   "Carrier_74_Status.7" AT %I4050.7 : Bool;   // CARRIER FAULT
   "Carrier_74_Status.8" AT %I4051.0 : Bool;   // CRASH DETECT TRIPPED
   "Carrier_74_Status.9" AT %I4051.1 : Bool;
   "Carrier_74_Status.10" AT %I4051.2 : Bool;
   "Carrier_74_Status.11" AT %I4051.3 : Bool;
   "Carrier_74_Status.12" AT %I4051.4 : Bool;
   "Carrier_74_Status.13" AT %I4051.5 : Bool;
   "Carrier_74_Status.14" AT %I4051.6 : Bool;
   "Carrier_74_Status.15" AT %I4051.7 : Bool;
   "Carrier_74_SDCFaultCode" AT %IW4052 : Word;   // SDC FAULT CODE
   "Carrier_74_CarrierPosition" AT %ID4054 : DWord;   // CARRIER POSITION
   "Carrier_74_CarrierNumber" AT %IW4058 : Word;   // CARRIER NUMBER
   "Carrier_74_G120DControlWord" AT %IW4060 : Word;   // G120D_STW1_CONTROL
   "Carrier_74_G120DControlWord.0" AT %I4060.0 : Bool;   // Bit_00_ON
   "Carrier_74_G120DControlWord.1" AT %I4060.1 : Bool;   // Bit_01_AUS2_INH
   "Carrier_74_G120DControlWord.2" AT %I4060.2 : Bool;   // Bit_02_AUS3_STOP
   "Carrier_74_G120DControlWord.3" AT %I4060.3 : Bool;   // Bit_03_EN
   "Carrier_74_G120DControlWord.4" AT %I4060.4 : Bool;   // Bit_04_EN_RAMP
   "Carrier_74_G120DControlWord.5" AT %I4060.5 : Bool;   // Bit_05_START_RAMP
   "Carrier_74_G120DControlWord.6" AT %I4060.6 : Bool;   // Bit_06_SETPOINT
   "Carrier_74_G120DControlWord.7" AT %I4060.7 : Bool;   // Bit_07_RESET
   "Carrier_74_G120DControlWord.8" AT %I4061.0 : Bool;   // Bit_08_JOG_R
   "Carrier_74_G120DControlWord.9" AT %I4061.1 : Bool;   // Bit_09_JOG_L
   "Carrier_74_G120DControlWord.10" AT %I4061.2 : Bool;   // Bit_10_CONTR_PLC
   "Carrier_74_G120DControlWord.11" AT %I4061.3 : Bool;   // Bit_11_REVERSE
   "Carrier_74_G120DControlWord.12" AT %I4061.4 : Bool;   // Bit_12_BRAKE_RELEASE
   "Carrier_74_G120DControlWord.13" AT %I4061.5 : Bool;   // Bit_13_DDS
   "Carrier_74_G120DControlWord.14" AT %I4061.6 : Bool;   // Bit_14_DO0
   "Carrier_74_G120DControlWord.15" AT %I4061.7 : Bool;   // Bit_15_DO1
   "Carrier_74_G120DStatusWord" AT %IW4062 : Word;   // G120D_ZSW1_STATUS
   "Carrier_74_G120DStatusWord.0" AT %I4062.0 : Bool;   // Bit_00_READY_RUN
   "Carrier_74_G120DStatusWord.1" AT %I4062.1 : Bool;   // Bit_01_READY_ON
   "Carrier_74_G120DStatusWord.2" AT %I4062.2 : Bool;   // Bit_02_ENABLE
   "Carrier_74_G120DStatusWord.3" AT %I4062.3 : Bool;   // Bit_03_FAULT
   "Carrier_74_G120DStatusWord.4" AT %I4062.4 : Bool;   // Bit_04_OFF2
   "Carrier_74_G120DStatusWord.5" AT %I4062.5 : Bool;   // Bit_05_OFF3
   "Carrier_74_G120DStatusWord.6" AT %I4062.6 : Bool;   // Bit_06_LOCK_OUT
   "Carrier_74_G120DStatusWord.7" AT %I4062.7 : Bool;   // Bit_07_WARN
   "Carrier_74_G120DStatusWord.8" AT %I4063.0 : Bool;   // Bit_08_NO_DEVIATION
   "Carrier_74_G120DStatusWord.9" AT %I4063.1 : Bool;   // Bit_09_CONTR_PLC
   "Carrier_74_G120DStatusWord.10" AT %I4063.2 : Bool;   // Bit_10_F_MAX
   "Carrier_74_G120DStatusWord.11" AT %I4063.3 : Bool;   // Bit_11_LIMIT_REACHED
   "Carrier_74_G120DStatusWord.12" AT %I4063.4 : Bool;   // Bit_12_BRAKE_OPEN
   "Carrier_74_G120DStatusWord.13" AT %I4063.5 : Bool;   // Bit_13_NO_OVERTEMP
   "Carrier_74_G120DStatusWord.14" AT %I4063.6 : Bool;   // Bit_14_CW_CCW
   "Carrier_74_G120DStatusWord.15" AT %I4063.7 : Bool;   // Bit_15_OVERL
   "Carrier_74_Slot2_Input" AT %IW4064 : Word;   // SLOT 2 INPUT WORD
   "Carrier_74_CrashDetectSW" AT %I4064.0 : Bool;   // CRASH DETECT SW
   "Carrier_74_SpareSafetyInput(2_1)" AT %I4064.1 : Bool;   // SPARE SAFETY INPUT
   "Carrier_74_SpareSafetyInput(2_2)" AT %I4064.2 : Bool;   // SPARE SAFETY INPUT
   "Carrier_74_SpareSafetyInput(2_3)" AT %I4064.3 : Bool;   // SPARE SAFETY INPUT
   "Carrier_74_SpareSafetyInput(2_4)" AT %I4064.4 : Bool;   // SPARE SAFETY INPUT
   "Carrier_74_SpareSafetyInput(2_5)" AT %I4064.5 : Bool;   // SPARE SAFETY INPUT
   "Carrier_74_SpareSafetyInput(2_6)" AT %I4064.6 : Bool;   // SPARE SAFETY INPUT
   "Carrier_74_SpareSafetyInput(2_7)" AT %I4064.7 : Bool;   // SPARE SAFETY INPUT
   "Carrier_74_Slot3_SafetyOutput" AT %IW4065 : Word;   // SLOT 3 SAFETY OUTPUT WORD
   "Carrier_74_Crash_Detect_OK" AT %I4065.0 : Bool;   // CARRIER CRASH DETECT
   "Carrier_74_SpareSafetyOutput(3_1)" AT %I4065.1 : Bool;   // SPARE SAFETY OUTPUT
   "Carrier_74_SpareSafetyOutput(3_2)" AT %I4065.2 : Bool;   // SPARE SAFETY OUTPUT
   "Carrier_74_SpareSafetyOutput(3_3)" AT %I4065.3 : Bool;   // SPARE SAFETY OUTPUT
   "Carrier_74_SpareSafetyOutput(3_4)" AT %I4065.4 : Bool;   // SPARE SAFETY OUTPUT
   "Carrier_74_SpareSafetyOutput(3_5)" AT %I4065.5 : Bool;   // SPARE SAFETY OUTPUT
   "Carrier_74_SpareSafetyOutput(3_6)" AT %I4065.6 : Bool;   // SPARE SAFETY OUTPUT
   "Carrier_74_SpareSafetyOutput(3_7)" AT %I4065.7 : Bool;   // SPARE SAFETY OUTPUT
   "Carrier_74_Slot4_Input" AT %IW4066 : Word;   // SLOT 4 INPUT WORD
   "Carrier_74_480VPowerOn_MDCB1" AT %I4066.0 : Bool;   // 480 VAC POWER ON MDCB 1
   "Carrier_74_SpareInput(4_1)" AT %I4066.1 : Bool;   // SPARE INPUT
   "Carrier_74_SpareInput(4_2)" AT %I4066.2 : Bool;   // SPARE INPUT
   "Carrier_74_SitopSelectStatus" AT %I4066.3 : Bool;   // SITOP SELECT STATUS
   "Carrier_74_DCsupplyOnPSCB2" AT %I4066.4 : Bool;   // DC SUPPLY ON PSCB 2
   "Carrier_74_SpareInput(4_5)" AT %I4066.5 : Bool;   // SPARE INPUT
   "Carrier_74_SpareInput(4_6)" AT %I4066.6 : Bool;   // SPARE INPUT
   "Carrier_74_SpareInput(4_7)" AT %I4066.7 : Bool;   // SPARE INPUT
   "Carrier_74_PB1_ProdHoldLH" AT %I4067.0 : Bool;   // PB 1 PRODUCTION HOLD LH
   "Carrier_74_PB2_ResetLH" AT %I4067.1 : Bool;   // PB 2 RESET LH
   "Carrier_74_PB3_ProdHoldRH" AT %I4067.2 : Bool;   // PB 3 PRODUCTION HOLD RH
   "Carrier_74_PB4_ResetRH" AT %I4067.3 : Bool;   // PB 4 RESET RH
   "Carrier_74_SpareInput(4_14)" AT %I4067.4 : Bool;   // SPARE INPUT
   "Carrier_74_SpareInput(4_15)" AT %I4067.5 : Bool;   // SPARE INPUT
   "Carrier_74_SpareInput(4_16)" AT %I4067.6 : Bool;   // SPARE INPUT
   "Carrier_74_SpareInput(4_17)" AT %I4067.7 : Bool;   // SPARE INPUT
   "Carrier_74_Slot5_Output" AT %IW4068 : Word;   // SLOT 5 OUTPUT WORD
   "Carrier_74_IRD400_HMI_24VDC_ENABLE" AT %I4068.0 : Bool;   // IRD 400 PANEL HMI 24V DC POWER
   "Carrier_74_FaultLight_LH" AT %I4068.1 : Bool;   // FAULT LIGHT LH
   "Carrier_74_RunLight_LH" AT %I4068.2 : Bool;   // RUN LIGHT LH
   "Carrier_74_FaultLight_RH" AT %I4068.3 : Bool;   // FAULT LIGHT RH
   "Carrier_74_RunLight_RH" AT %I4068.4 : Bool;   // RUN LIGHT RH
   "Carrier_74_SpareOutput(5_5)" AT %I4068.5 : Bool;   // SPARE OUTPUT
   "Carrier_74_SpareOutput(5_6)" AT %I4068.6 : Bool;   // SPARE OUTPUT
   "Carrier_74_SpareOutput(5_7)" AT %I4068.7 : Bool;   // SPARE OUTPUT
   "Carrier_74_ActualSpeed" AT %IW4070 : Word;   // ACTUAL SPEED
   "Carrier_74_CarrierDriveAlarm" AT %IW4072 : Word;   // CARRIER DRIVE ALARM
   "Carrier_74_CarrierDriveWarning" AT %IW4074 : Word;   // CARRIER DRIVE WARNING
   "Carrier_75_Status" AT %IW4100 : Word;   // CARRIER STATUS WORD
   "Carrier_75_Status.0" AT %I4100.0 : Bool;   // HEARTBEAT
   "Carrier_75_Status.1" AT %I4100.1 : Bool;   // MANUAL
   "Carrier_75_Status.2" AT %I4100.2 : Bool;   // IN_AUTO
   "Carrier_75_Status.3" AT %I4100.3 : Bool;   // POSITIONING_COMPLETE
   "Carrier_75_Status.4" AT %I4100.4 : Bool;   // PRODUCTION HOLD
   "Carrier_75_Status.5" AT %I4100.5 : Bool;   // CARRIER MOVING FORWARD
   "Carrier_75_Status.6" AT %I4100.6 : Bool;   // CARRIER MOVING REVERSE
   "Carrier_75_Status.7" AT %I4100.7 : Bool;   // CARRIER FAULT
   "Carrier_75_Status.8" AT %I4101.0 : Bool;   // CRASH DETECT TRIPPED
   "Carrier_75_Status.9" AT %I4101.1 : Bool;
   "Carrier_75_Status.10" AT %I4101.2 : Bool;
   "Carrier_75_Status.11" AT %I4101.3 : Bool;
   "Carrier_75_Status.12" AT %I4101.4 : Bool;
   "Carrier_75_Status.13" AT %I4101.5 : Bool;
   "Carrier_75_Status.14" AT %I4101.6 : Bool;
   "Carrier_75_Status.15" AT %I4101.7 : Bool;
   "Carrier_75_SDCFaultCode" AT %IW4102 : Word;   // SDC FAULT CODE
   "Carrier_75_CarrierPosition" AT %ID4104 : DWord;   // CARRIER POSITION
   "Carrier_75_CarrierNumber" AT %IW4108 : Word;   // CARRIER NUMBER
   "Carrier_75_G120DControlWord" AT %IW4110 : Word;   // G120D_STW1_CONTROL
   "Carrier_75_G120DControlWord.0" AT %I4110.0 : Bool;   // Bit_00_ON
   "Carrier_75_G120DControlWord.1" AT %I4110.1 : Bool;   // Bit_01_AUS2_INH
   "Carrier_75_G120DControlWord.2" AT %I4110.2 : Bool;   // Bit_02_AUS3_STOP
   "Carrier_75_G120DControlWord.3" AT %I4110.3 : Bool;   // Bit_03_EN
   "Carrier_75_G120DControlWord.4" AT %I4110.4 : Bool;   // Bit_04_EN_RAMP
   "Carrier_75_G120DControlWord.5" AT %I4110.5 : Bool;   // Bit_05_START_RAMP
   "Carrier_75_G120DControlWord.6" AT %I4110.6 : Bool;   // Bit_06_SETPOINT
   "Carrier_75_G120DControlWord.7" AT %I4110.7 : Bool;   // Bit_07_RESET
   "Carrier_75_G120DControlWord.8" AT %I4111.0 : Bool;   // Bit_08_JOG_R
   "Carrier_75_G120DControlWord.9" AT %I4111.1 : Bool;   // Bit_09_JOG_L
   "Carrier_75_G120DControlWord.10" AT %I4111.2 : Bool;   // Bit_10_CONTR_PLC
   "Carrier_75_G120DControlWord.11" AT %I4111.3 : Bool;   // Bit_11_REVERSE
   "Carrier_75_G120DControlWord.12" AT %I4111.4 : Bool;   // Bit_12_BRAKE_RELEASE
   "Carrier_75_G120DControlWord.13" AT %I4111.5 : Bool;   // Bit_13_DDS
   "Carrier_75_G120DControlWord.14" AT %I4111.6 : Bool;   // Bit_14_DO0
   "Carrier_75_G120DControlWord.15" AT %I4111.7 : Bool;   // Bit_15_DO1
   "Carrier_75_G120DStatusWord" AT %IW4112 : Word;   // G120D_ZSW1_STATUS
   "Carrier_75_G120DStatusWord.0" AT %I4112.0 : Bool;   // Bit_00_READY_RUN
   "Carrier_75_G120DStatusWord.1" AT %I4112.1 : Bool;   // Bit_01_READY_ON
   "Carrier_75_G120DStatusWord.2" AT %I4112.2 : Bool;   // Bit_02_ENABLE
   "Carrier_75_G120DStatusWord.3" AT %I4112.3 : Bool;   // Bit_03_FAULT
   "Carrier_75_G120DStatusWord.4" AT %I4112.4 : Bool;   // Bit_04_OFF2
   "Carrier_75_G120DStatusWord.5" AT %I4112.5 : Bool;   // Bit_05_OFF3
   "Carrier_75_G120DStatusWord.6" AT %I4112.6 : Bool;   // Bit_06_LOCK_OUT
   "Carrier_75_G120DStatusWord.7" AT %I4112.7 : Bool;   // Bit_07_WARN
   "Carrier_75_G120DStatusWord.8" AT %I4113.0 : Bool;   // Bit_08_NO_DEVIATION
   "Carrier_75_G120DStatusWord.9" AT %I4113.1 : Bool;   // Bit_09_CONTR_PLC
   "Carrier_75_G120DStatusWord.10" AT %I4113.2 : Bool;   // Bit_10_F_MAX
   "Carrier_75_G120DStatusWord.11" AT %I4113.3 : Bool;   // Bit_11_LIMIT_REACHED
   "Carrier_75_G120DStatusWord.12" AT %I4113.4 : Bool;   // Bit_12_BRAKE_OPEN
   "Carrier_75_G120DStatusWord.13" AT %I4113.5 : Bool;   // Bit_13_NO_OVERTEMP
   "Carrier_75_G120DStatusWord.14" AT %I4113.6 : Bool;   // Bit_14_CW_CCW
   "Carrier_75_G120DStatusWord.15" AT %I4113.7 : Bool;   // Bit_15_OVERL
   "Carrier_75_Slot2_Input" AT %IW4114 : Word;   // SLOT 2 INPUT WORD
   "Carrier_75_CrashDetectSW" AT %I4114.0 : Bool;   // CRASH DETECT SW
   "Carrier_75_SpareSafetyInput(2_1)" AT %I4114.1 : Bool;   // SPARE SAFETY INPUT
   "Carrier_75_SpareSafetyInput(2_2)" AT %I4114.2 : Bool;   // SPARE SAFETY INPUT
   "Carrier_75_SpareSafetyInput(2_3)" AT %I4114.3 : Bool;   // SPARE SAFETY INPUT
   "Carrier_75_SpareSafetyInput(2_4)" AT %I4114.4 : Bool;   // SPARE SAFETY INPUT
   "Carrier_75_SpareSafetyInput(2_5)" AT %I4114.5 : Bool;   // SPARE SAFETY INPUT
   "Carrier_75_SpareSafetyInput(2_6)" AT %I4114.6 : Bool;   // SPARE SAFETY INPUT
   "Carrier_75_SpareSafetyInput(2_7)" AT %I4114.7 : Bool;   // SPARE SAFETY INPUT
   "Carrier_75_Slot3_SafetyOutput" AT %IW4115 : Word;   // SLOT 3 SAFETY OUTPUT WORD
   "Carrier_75_Crash_Detect_OK" AT %I4115.0 : Bool;   // CARRIER CRASH DETECT
   "Carrier_75_SpareSafetyOutput(3_1)" AT %I4115.1 : Bool;   // SPARE SAFETY OUTPUT
   "Carrier_75_SpareSafetyOutput(3_2)" AT %I4115.2 : Bool;   // SPARE SAFETY OUTPUT
   "Carrier_75_SpareSafetyOutput(3_3)" AT %I4115.3 : Bool;   // SPARE SAFETY OUTPUT
   "Carrier_75_SpareSafetyOutput(3_4)" AT %I4115.4 : Bool;   // SPARE SAFETY OUTPUT
   "Carrier_75_SpareSafetyOutput(3_5)" AT %I4115.5 : Bool;   // SPARE SAFETY OUTPUT
   "Carrier_75_SpareSafetyOutput(3_6)" AT %I4115.6 : Bool;   // SPARE SAFETY OUTPUT
   "Carrier_75_SpareSafetyOutput(3_7)" AT %I4115.7 : Bool;   // SPARE SAFETY OUTPUT
   "Carrier_75_Slot4_Input" AT %IW4116 : Word;   // SLOT 4 INPUT WORD
   "Carrier_75_480VPowerOn_MDCB1" AT %I4116.0 : Bool;   // 480 VAC POWER ON MDCB 1
   "Carrier_75_SpareInput(4_1)" AT %I4116.1 : Bool;   // SPARE INPUT
   "Carrier_75_SpareInput(4_2)" AT %I4116.2 : Bool;   // SPARE INPUT
   "Carrier_75_SitopSelectStatus" AT %I4116.3 : Bool;   // SITOP SELECT STATUS
   "Carrier_75_DCsupplyOnPSCB2" AT %I4116.4 : Bool;   // DC SUPPLY ON PSCB 2
   "Carrier_75_SpareInput(4_5)" AT %I4116.5 : Bool;   // SPARE INPUT
   "Carrier_75_SpareInput(4_6)" AT %I4116.6 : Bool;   // SPARE INPUT
   "Carrier_75_SpareInput(4_7)" AT %I4116.7 : Bool;   // SPARE INPUT
   "Carrier_75_PB1_ProdHoldLH" AT %I4117.0 : Bool;   // PB 1 PRODUCTION HOLD LH
   "Carrier_75_PB2_ResetLH" AT %I4117.1 : Bool;   // PB 2 RESET LH
   "Carrier_75_PB3_ProdHoldRH" AT %I4117.2 : Bool;   // PB 3 PRODUCTION HOLD RH
   "Carrier_75_PB4_ResetRH" AT %I4117.3 : Bool;   // PB 4 RESET RH
   "Carrier_75_SpareInput(4_14)" AT %I4117.4 : Bool;   // SPARE INPUT
   "Carrier_75_SpareInput(4_15)" AT %I4117.5 : Bool;   // SPARE INPUT
   "Carrier_75_SpareInput(4_16)" AT %I4117.6 : Bool;   // SPARE INPUT
   "Carrier_75_SpareInput(4_17)" AT %I4117.7 : Bool;   // SPARE INPUT
   "Carrier_75_Slot5_Output" AT %IW4118 : Word;   // SLOT 5 OUTPUT WORD
   "Carrier_75_IRD400_HMI_24VDC_ENABLE" AT %I4118.0 : Bool;   // IRD 400 PANEL HMI 24V DC POWER
   "Carrier_75_FaultLight_LH" AT %I4118.1 : Bool;   // FAULT LIGHT LH
   "Carrier_75_RunLight_LH" AT %I4118.2 : Bool;   // RUN LIGHT LH
   "Carrier_75_FaultLight_RH" AT %I4118.3 : Bool;   // FAULT LIGHT RH
   "Carrier_75_RunLight_RH" AT %I4118.4 : Bool;   // RUN LIGHT RH
   "Carrier_75_SpareOutput(5_5)" AT %I4118.5 : Bool;   // SPARE OUTPUT
   "Carrier_75_SpareOutput(5_6)" AT %I4118.6 : Bool;   // SPARE OUTPUT
   "Carrier_75_SpareOutput(5_7)" AT %I4118.7 : Bool;   // SPARE OUTPUT
   "Carrier_75_ActualSpeed" AT %IW4120 : Word;   // ACTUAL SPEED
   "Carrier_75_CarrierDriveAlarm" AT %IW4122 : Word;   // CARRIER DRIVE ALARM
   "Carrier_75_CarrierDriveWarning" AT %IW4124 : Word;   // CARRIER DRIVE WARNING
   "Carrier_76_Status" AT %IW4150 : Word;   // CARRIER STATUS WORD
   "Carrier_76_Status.0" AT %I4150.0 : Bool;   // HEARTBEAT
   "Carrier_76_Status.1" AT %I4150.1 : Bool;   // MANUAL
   "Carrier_76_Status.2" AT %I4150.2 : Bool;   // IN_AUTO
   "Carrier_76_Status.3" AT %I4150.3 : Bool;   // POSITIONING_COMPLETE
   "Carrier_76_Status.4" AT %I4150.4 : Bool;   // PRODUCTION HOLD
   "Carrier_76_Status.5" AT %I4150.5 : Bool;   // CARRIER MOVING FORWARD
   "Carrier_76_Status.6" AT %I4150.6 : Bool;   // CARRIER MOVING REVERSE
   "Carrier_76_Status.7" AT %I4150.7 : Bool;   // CARRIER FAULT
   "Carrier_76_Status.8" AT %I4151.0 : Bool;   // CRASH DETECT TRIPPED
   "Carrier_76_Status.9" AT %I4151.1 : Bool;
   "Carrier_76_Status.10" AT %I4151.2 : Bool;
   "Carrier_76_Status.11" AT %I4151.3 : Bool;
   "Carrier_76_Status.12" AT %I4151.4 : Bool;
   "Carrier_76_Status.13" AT %I4151.5 : Bool;
   "Carrier_76_Status.14" AT %I4151.6 : Bool;
   "Carrier_76_Status.15" AT %I4151.7 : Bool;
   "Carrier_76_SDCFaultCode" AT %IW4152 : Word;   // SDC FAULT CODE
   "Carrier_76_CarrierPosition" AT %ID4154 : DWord;   // CARRIER POSITION
   "Carrier_76_CarrierNumber" AT %IW4158 : Word;   // CARRIER NUMBER
   "Carrier_76_G120DControlWord" AT %IW4160 : Word;   // G120D_STW1_CONTROL
   "Carrier_76_G120DControlWord.0" AT %I4160.0 : Bool;   // Bit_00_ON
   "Carrier_76_G120DControlWord.1" AT %I4160.1 : Bool;   // Bit_01_AUS2_INH
   "Carrier_76_G120DControlWord.2" AT %I4160.2 : Bool;   // Bit_02_AUS3_STOP
   "Carrier_76_G120DControlWord.3" AT %I4160.3 : Bool;   // Bit_03_EN
   "Carrier_76_G120DControlWord.4" AT %I4160.4 : Bool;   // Bit_04_EN_RAMP
   "Carrier_76_G120DControlWord.5" AT %I4160.5 : Bool;   // Bit_05_START_RAMP
   "Carrier_76_G120DControlWord.6" AT %I4160.6 : Bool;   // Bit_06_SETPOINT
   "Carrier_76_G120DControlWord.7" AT %I4160.7 : Bool;   // Bit_07_RESET
   "Carrier_76_G120DControlWord.8" AT %I4161.0 : Bool;   // Bit_08_JOG_R
   "Carrier_76_G120DControlWord.9" AT %I4161.1 : Bool;   // Bit_09_JOG_L
   "Carrier_76_G120DControlWord.10" AT %I4161.2 : Bool;   // Bit_10_CONTR_PLC
   "Carrier_76_G120DControlWord.11" AT %I4161.3 : Bool;   // Bit_11_REVERSE
   "Carrier_76_G120DControlWord.12" AT %I4161.4 : Bool;   // Bit_12_BRAKE_RELEASE
   "Carrier_76_G120DControlWord.13" AT %I4161.5 : Bool;   // Bit_13_DDS
   "Carrier_76_G120DControlWord.14" AT %I4161.6 : Bool;   // Bit_14_DO0
   "Carrier_76_G120DControlWord.15" AT %I4161.7 : Bool;   // Bit_15_DO1
   "Carrier_76_G120DStatusWord" AT %IW4162 : Word;   // G120D_ZSW1_STATUS
   "Carrier_76_G120DStatusWord.0" AT %I4162.0 : Bool;   // Bit_00_READY_RUN
   "Carrier_76_G120DStatusWord.1" AT %I4162.1 : Bool;   // Bit_01_READY_ON
   "Carrier_76_G120DStatusWord.2" AT %I4162.2 : Bool;   // Bit_02_ENABLE
   "Carrier_76_G120DStatusWord.3" AT %I4162.3 : Bool;   // Bit_03_FAULT
   "Carrier_76_G120DStatusWord.4" AT %I4162.4 : Bool;   // Bit_04_OFF2
   "Carrier_76_G120DStatusWord.5" AT %I4162.5 : Bool;   // Bit_05_OFF3
   "Carrier_76_G120DStatusWord.6" AT %I4162.6 : Bool;   // Bit_06_LOCK_OUT
   "Carrier_76_G120DStatusWord.7" AT %I4162.7 : Bool;   // Bit_07_WARN
   "Carrier_76_G120DStatusWord.8" AT %I4163.0 : Bool;   // Bit_08_NO_DEVIATION
   "Carrier_76_G120DStatusWord.9" AT %I4163.1 : Bool;   // Bit_09_CONTR_PLC
   "Carrier_76_G120DStatusWord.10" AT %I4163.2 : Bool;   // Bit_10_F_MAX
   "Carrier_76_G120DStatusWord.11" AT %I4163.3 : Bool;   // Bit_11_LIMIT_REACHED
   "Carrier_76_G120DStatusWord.12" AT %I4163.4 : Bool;   // Bit_12_BRAKE_OPEN
   "Carrier_76_G120DStatusWord.13" AT %I4163.5 : Bool;   // Bit_13_NO_OVERTEMP
   "Carrier_76_G120DStatusWord.14" AT %I4163.6 : Bool;   // Bit_14_CW_CCW
   "Carrier_76_G120DStatusWord.15" AT %I4163.7 : Bool;   // Bit_15_OVERL
   "Carrier_76_Slot2_Input" AT %IW4164 : Word;   // SLOT 2 INPUT WORD
   "Carrier_76_CrashDetectSW" AT %I4164.0 : Bool;   // CRASH DETECT SW
   "Carrier_76_SpareSafetyInput(2_1)" AT %I4164.1 : Bool;   // SPARE SAFETY INPUT
   "Carrier_76_SpareSafetyInput(2_2)" AT %I4164.2 : Bool;   // SPARE SAFETY INPUT
   "Carrier_76_SpareSafetyInput(2_3)" AT %I4164.3 : Bool;   // SPARE SAFETY INPUT
   "Carrier_76_SpareSafetyInput(2_4)" AT %I4164.4 : Bool;   // SPARE SAFETY INPUT
   "Carrier_76_SpareSafetyInput(2_5)" AT %I4164.5 : Bool;   // SPARE SAFETY INPUT
   "Carrier_76_SpareSafetyInput(2_6)" AT %I4164.6 : Bool;   // SPARE SAFETY INPUT
   "Carrier_76_SpareSafetyInput(2_7)" AT %I4164.7 : Bool;   // SPARE SAFETY INPUT
   "Carrier_76_Slot3_SafetyOutput" AT %IW4165 : Word;   // SLOT 3 SAFETY OUTPUT WORD
   "Carrier_76_Crash_Detect_OK" AT %I4165.0 : Bool;   // CARRIER CRASH DETECT
   "Carrier_76_SpareSafetyOutput(3_1)" AT %I4165.1 : Bool;   // SPARE SAFETY OUTPUT
   "Carrier_76_SpareSafetyOutput(3_2)" AT %I4165.2 : Bool;   // SPARE SAFETY OUTPUT
   "Carrier_76_SpareSafetyOutput(3_3)" AT %I4165.3 : Bool;   // SPARE SAFETY OUTPUT
   "Carrier_76_SpareSafetyOutput(3_4)" AT %I4165.4 : Bool;   // SPARE SAFETY OUTPUT
   "Carrier_76_SpareSafetyOutput(3_5)" AT %I4165.5 : Bool;   // SPARE SAFETY OUTPUT
   "Carrier_76_SpareSafetyOutput(3_6)" AT %I4165.6 : Bool;   // SPARE SAFETY OUTPUT
   "Carrier_76_SpareSafetyOutput(3_7)" AT %I4165.7 : Bool;   // SPARE SAFETY OUTPUT
   "Carrier_76_Slot4_Input" AT %IW4166 : Word;   // SLOT 4 INPUT WORD
   "Carrier_76_480VPowerOn_MDCB1" AT %I4166.0 : Bool;   // 480 VAC POWER ON MDCB 1
   "Carrier_76_SpareInput(4_1)" AT %I4166.1 : Bool;   // SPARE INPUT
   "Carrier_76_SpareInput(4_2)" AT %I4166.2 : Bool;   // SPARE INPUT
   "Carrier_76_SitopSelectStatus" AT %I4166.3 : Bool;   // SITOP SELECT STATUS
   "Carrier_76_DCsupplyOnPSCB2" AT %I4166.4 : Bool;   // DC SUPPLY ON PSCB 2
   "Carrier_76_SpareInput(4_5)" AT %I4166.5 : Bool;   // SPARE INPUT
   "Carrier_76_SpareInput(4_6)" AT %I4166.6 : Bool;   // SPARE INPUT
   "Carrier_76_SpareInput(4_7)" AT %I4166.7 : Bool;   // SPARE INPUT
   "Carrier_76_PB1_ProdHoldLH" AT %I4167.0 : Bool;   // PB 1 PRODUCTION HOLD LH
   "Carrier_76_PB2_ResetLH" AT %I4167.1 : Bool;   // PB 2 RESET LH
   "Carrier_76_PB3_ProdHoldRH" AT %I4167.2 : Bool;   // PB 3 PRODUCTION HOLD RH
   "Carrier_76_PB4_ResetRH" AT %I4167.3 : Bool;   // PB 4 RESET RH
   "Carrier_76_SpareInput(4_14)" AT %I4167.4 : Bool;   // SPARE INPUT
   "Carrier_76_SpareInput(4_15)" AT %I4167.5 : Bool;   // SPARE INPUT
   "Carrier_76_SpareInput(4_16)" AT %I4167.6 : Bool;   // SPARE INPUT
   "Carrier_76_SpareInput(4_17)" AT %I4167.7 : Bool;   // SPARE INPUT
   "Carrier_76_Slot5_Output" AT %IW4168 : Word;   // SLOT 5 OUTPUT WORD
   "Carrier_76_IRD400_HMI_24VDC_ENABLE" AT %I4168.0 : Bool;   // IRD 400 PANEL HMI 24V DC POWER
   "Carrier_76_FaultLight_LH" AT %I4168.1 : Bool;   // FAULT LIGHT LH
   "Carrier_76_RunLight_LH" AT %I4168.2 : Bool;   // RUN LIGHT LH
   "Carrier_76_FaultLight_RH" AT %I4168.3 : Bool;   // FAULT LIGHT RH
   "Carrier_76_RunLight_RH" AT %I4168.4 : Bool;   // RUN LIGHT RH
   "Carrier_76_SpareOutput(5_5)" AT %I4168.5 : Bool;   // SPARE OUTPUT
   "Carrier_76_SpareOutput(5_6)" AT %I4168.6 : Bool;   // SPARE OUTPUT
   "Carrier_76_SpareOutput(5_7)" AT %I4168.7 : Bool;   // SPARE OUTPUT
   "Carrier_76_ActualSpeed" AT %IW4170 : Word;   // ACTUAL SPEED
   "Carrier_76_CarrierDriveAlarm" AT %IW4172 : Word;   // CARRIER DRIVE ALARM
   "Carrier_76_CarrierDriveWarning" AT %IW4174 : Word;   // CARRIER DRIVE WARNING
   "Carrier_77_Status" AT %IW4200 : Word;   // CARRIER STATUS WORD
   "Carrier_77_Status.0" AT %I4200.0 : Bool;   // HEARTBEAT
   "Carrier_77_Status.1" AT %I4200.1 : Bool;   // MANUAL
   "Carrier_77_Status.2" AT %I4200.2 : Bool;   // IN_AUTO
   "Carrier_77_Status.3" AT %I4200.3 : Bool;   // POSITIONING_COMPLETE
   "Carrier_77_Status.4" AT %I4200.4 : Bool;   // PRODUCTION HOLD
   "Carrier_77_Status.5" AT %I4200.5 : Bool;   // CARRIER MOVING FORWARD
   "Carrier_77_Status.6" AT %I4200.6 : Bool;   // CARRIER MOVING REVERSE
   "Carrier_77_Status.7" AT %I4200.7 : Bool;   // CARRIER FAULT
   "Carrier_77_Status.8" AT %I4201.0 : Bool;   // CRASH DETECT TRIPPED
   "Carrier_77_Status.9" AT %I4201.1 : Bool;
   "Carrier_77_Status.10" AT %I4201.2 : Bool;
   "Carrier_77_Status.11" AT %I4201.3 : Bool;
   "Carrier_77_Status.12" AT %I4201.4 : Bool;
   "Carrier_77_Status.13" AT %I4201.5 : Bool;
   "Carrier_77_Status.14" AT %I4201.6 : Bool;
   "Carrier_77_Status.15" AT %I4201.7 : Bool;
   "Carrier_77_SDCFaultCode" AT %IW4202 : Word;   // SDC FAULT CODE
   "Carrier_77_CarrierPosition" AT %ID4204 : DWord;   // CARRIER POSITION
   "Carrier_77_CarrierNumber" AT %IW4208 : Word;   // CARRIER NUMBER
   "Carrier_77_G120DControlWord" AT %IW4210 : Word;   // G120D_STW1_CONTROL
   "Carrier_77_G120DControlWord.0" AT %I4210.0 : Bool;   // Bit_00_ON
   "Carrier_77_G120DControlWord.1" AT %I4210.1 : Bool;   // Bit_01_AUS2_INH
   "Carrier_77_G120DControlWord.2" AT %I4210.2 : Bool;   // Bit_02_AUS3_STOP
   "Carrier_77_G120DControlWord.3" AT %I4210.3 : Bool;   // Bit_03_EN
   "Carrier_77_G120DControlWord.4" AT %I4210.4 : Bool;   // Bit_04_EN_RAMP
   "Carrier_77_G120DControlWord.5" AT %I4210.5 : Bool;   // Bit_05_START_RAMP
   "Carrier_77_G120DControlWord.6" AT %I4210.6 : Bool;   // Bit_06_SETPOINT
   "Carrier_77_G120DControlWord.7" AT %I4210.7 : Bool;   // Bit_07_RESET
   "Carrier_77_G120DControlWord.8" AT %I4211.0 : Bool;   // Bit_08_JOG_R
   "Carrier_77_G120DControlWord.9" AT %I4211.1 : Bool;   // Bit_09_JOG_L
   "Carrier_77_G120DControlWord.10" AT %I4211.2 : Bool;   // Bit_10_CONTR_PLC
   "Carrier_77_G120DControlWord.11" AT %I4211.3 : Bool;   // Bit_11_REVERSE
   "Carrier_77_G120DControlWord.12" AT %I4211.4 : Bool;   // Bit_12_BRAKE_RELEASE
   "Carrier_77_G120DControlWord.13" AT %I4211.5 : Bool;   // Bit_13_DDS
   "Carrier_77_G120DControlWord.14" AT %I4211.6 : Bool;   // Bit_14_DO0
   "Carrier_77_G120DControlWord.15" AT %I4211.7 : Bool;   // Bit_15_DO1
   "Carrier_77_G120DStatusWord" AT %IW4212 : Word;   // G120D_ZSW1_STATUS
   "Carrier_77_G120DStatusWord.0" AT %I4212.0 : Bool;   // Bit_00_READY_RUN
   "Carrier_77_G120DStatusWord.1" AT %I4212.1 : Bool;   // Bit_01_READY_ON
   "Carrier_77_G120DStatusWord.2" AT %I4212.2 : Bool;   // Bit_02_ENABLE
   "Carrier_77_G120DStatusWord.3" AT %I4212.3 : Bool;   // Bit_03_FAULT
   "Carrier_77_G120DStatusWord.4" AT %I4212.4 : Bool;   // Bit_04_OFF2
   "Carrier_77_G120DStatusWord.5" AT %I4212.5 : Bool;   // Bit_05_OFF3
   "Carrier_77_G120DStatusWord.6" AT %I4212.6 : Bool;   // Bit_06_LOCK_OUT
   "Carrier_77_G120DStatusWord.7" AT %I4212.7 : Bool;   // Bit_07_WARN
   "Carrier_77_G120DStatusWord.8" AT %I4213.0 : Bool;   // Bit_08_NO_DEVIATION
   "Carrier_77_G120DStatusWord.9" AT %I4213.1 : Bool;   // Bit_09_CONTR_PLC
   "Carrier_77_G120DStatusWord.10" AT %I4213.2 : Bool;   // Bit_10_F_MAX
   "Carrier_77_G120DStatusWord.11" AT %I4213.3 : Bool;   // Bit_11_LIMIT_REACHED
   "Carrier_77_G120DStatusWord.12" AT %I4213.4 : Bool;   // Bit_12_BRAKE_OPEN
   "Carrier_77_G120DStatusWord.13" AT %I4213.5 : Bool;   // Bit_13_NO_OVERTEMP
   "Carrier_77_G120DStatusWord.14" AT %I4213.6 : Bool;   // Bit_14_CW_CCW
   "Carrier_77_G120DStatusWord.15" AT %I4213.7 : Bool;   // Bit_15_OVERL
   "Carrier_77_Slot2_Input" AT %IW4214 : Word;   // SLOT 2 INPUT WORD
   "Carrier_77_CrashDetectSW" AT %I4214.0 : Bool;   // CRASH DETECT SW
   "Carrier_77_SpareSafetyInput(2_1)" AT %I4214.1 : Bool;   // SPARE SAFETY INPUT
   "Carrier_77_SpareSafetyInput(2_2)" AT %I4214.2 : Bool;   // SPARE SAFETY INPUT
   "Carrier_77_SpareSafetyInput(2_3)" AT %I4214.3 : Bool;   // SPARE SAFETY INPUT
   "Carrier_77_SpareSafetyInput(2_4)" AT %I4214.4 : Bool;   // SPARE SAFETY INPUT
   "Carrier_77_SpareSafetyInput(2_5)" AT %I4214.5 : Bool;   // SPARE SAFETY INPUT
   "Carrier_77_SpareSafetyInput(2_6)" AT %I4214.6 : Bool;   // SPARE SAFETY INPUT
   "Carrier_77_SpareSafetyInput(2_7)" AT %I4214.7 : Bool;   // SPARE SAFETY INPUT
   "Carrier_77_Slot3_SafetyOutput" AT %IW4215 : Word;   // SLOT 3 SAFETY OUTPUT WORD
   "Carrier_77_Crash_Detect_OK" AT %I4215.0 : Bool;   // CARRIER CRASH DETECT
   "Carrier_77_SpareSafetyOutput(3_1)" AT %I4215.1 : Bool;   // SPARE SAFETY OUTPUT
   "Carrier_77_SpareSafetyOutput(3_2)" AT %I4215.2 : Bool;   // SPARE SAFETY OUTPUT
   "Carrier_77_SpareSafetyOutput(3_3)" AT %I4215.3 : Bool;   // SPARE SAFETY OUTPUT
   "Carrier_77_SpareSafetyOutput(3_4)" AT %I4215.4 : Bool;   // SPARE SAFETY OUTPUT
   "Carrier_77_SpareSafetyOutput(3_5)" AT %I4215.5 : Bool;   // SPARE SAFETY OUTPUT
   "Carrier_77_SpareSafetyOutput(3_6)" AT %I4215.6 : Bool;   // SPARE SAFETY OUTPUT
   "Carrier_77_SpareSafetyOutput(3_7)" AT %I4215.7 : Bool;   // SPARE SAFETY OUTPUT
   "Carrier_77_Slot4_Input" AT %IW4216 : Word;   // SLOT 4 INPUT WORD
   "Carrier_77_480VPowerOn_MDCB1" AT %I4216.0 : Bool;   // 480 VAC POWER ON MDCB 1
   "Carrier_77_SpareInput(4_1)" AT %I4216.1 : Bool;   // SPARE INPUT
   "Carrier_77_SpareInput(4_2)" AT %I4216.2 : Bool;   // SPARE INPUT
   "Carrier_77_SitopSelectStatus" AT %I4216.3 : Bool;   // SITOP SELECT STATUS
   "Carrier_77_DCsupplyOnPSCB2" AT %I4216.4 : Bool;   // DC SUPPLY ON PSCB 2
   "Carrier_77_SpareInput(4_5)" AT %I4216.5 : Bool;   // SPARE INPUT
   "Carrier_77_SpareInput(4_6)" AT %I4216.6 : Bool;   // SPARE INPUT
   "Carrier_77_SpareInput(4_7)" AT %I4216.7 : Bool;   // SPARE INPUT
   "Carrier_77_PB1_ProdHoldLH" AT %I4217.0 : Bool;   // PB 1 PRODUCTION HOLD LH
   "Carrier_77_PB2_ResetLH" AT %I4217.1 : Bool;   // PB 2 RESET LH
   "Carrier_77_PB3_ProdHoldRH" AT %I4217.2 : Bool;   // PB 3 PRODUCTION HOLD RH
   "Carrier_77_PB4_ResetRH" AT %I4217.3 : Bool;   // PB 4 RESET RH
   "Carrier_77_SpareInput(4_14)" AT %I4217.4 : Bool;   // SPARE INPUT
   "Carrier_77_SpareInput(4_15)" AT %I4217.5 : Bool;   // SPARE INPUT
   "Carrier_77_SpareInput(4_16)" AT %I4217.6 : Bool;   // SPARE INPUT
   "Carrier_77_SpareInput(4_17)" AT %I4217.7 : Bool;   // SPARE INPUT
   "Carrier_77_Slot5_Output" AT %IW4218 : Word;   // SLOT 5 OUTPUT WORD
   "Carrier_77_IRD400_HMI_24VDC_ENABLE" AT %I4218.0 : Bool;   // IRD 400 PANEL HMI 24V DC POWER
   "Carrier_77_FaultLight_LH" AT %I4218.1 : Bool;   // FAULT LIGHT LH
   "Carrier_77_RunLight_LH" AT %I4218.2 : Bool;   // RUN LIGHT LH
   "Carrier_77_FaultLight_RH" AT %I4218.3 : Bool;   // FAULT LIGHT RH
   "Carrier_77_RunLight_RH" AT %I4218.4 : Bool;   // RUN LIGHT RH
   "Carrier_77_SpareOutput(5_5)" AT %I4218.5 : Bool;   // SPARE OUTPUT
   "Carrier_77_SpareOutput(5_6)" AT %I4218.6 : Bool;   // SPARE OUTPUT
   "Carrier_77_SpareOutput(5_7)" AT %I4218.7 : Bool;   // SPARE OUTPUT
   "Carrier_77_ActualSpeed" AT %IW4220 : Word;   // ACTUAL SPEED
   "Carrier_77_CarrierDriveAlarm" AT %IW4222 : Word;   // CARRIER DRIVE ALARM
   "Carrier_77_CarrierDriveWarning" AT %IW4224 : Word;   // CARRIER DRIVE WARNING
   "Carrier_78_Status" AT %IW4250 : Word;   // CARRIER STATUS WORD
   "Carrier_78_Status.0" AT %I4250.0 : Bool;   // HEARTBEAT
   "Carrier_78_Status.1" AT %I4250.1 : Bool;   // MANUAL
   "Carrier_78_Status.2" AT %I4250.2 : Bool;   // IN_AUTO
   "Carrier_78_Status.3" AT %I4250.3 : Bool;   // POSITIONING_COMPLETE
   "Carrier_78_Status.4" AT %I4250.4 : Bool;   // PRODUCTION HOLD
   "Carrier_78_Status.5" AT %I4250.5 : Bool;   // CARRIER MOVING FORWARD
   "Carrier_78_Status.6" AT %I4250.6 : Bool;   // CARRIER MOVING REVERSE
   "Carrier_78_Status.7" AT %I4250.7 : Bool;   // CARRIER FAULT
   "Carrier_78_Status.8" AT %I4251.0 : Bool;   // CRASH DETECT TRIPPED
   "Carrier_78_Status.9" AT %I4251.1 : Bool;
   "Carrier_78_Status.10" AT %I4251.2 : Bool;
   "Carrier_78_Status.11" AT %I4251.3 : Bool;
   "Carrier_78_Status.12" AT %I4251.4 : Bool;
   "Carrier_78_Status.13" AT %I4251.5 : Bool;
   "Carrier_78_Status.14" AT %I4251.6 : Bool;
   "Carrier_78_Status.15" AT %I4251.7 : Bool;
   "Carrier_78_SDCFaultCode" AT %IW4252 : Word;   // SDC FAULT CODE
   "Carrier_78_CarrierPosition" AT %ID4254 : DWord;   // CARRIER POSITION
   "Carrier_78_CarrierNumber" AT %IW4258 : Word;   // CARRIER NUMBER
   "Carrier_78_G120DControlWord" AT %IW4260 : Word;   // G120D_STW1_CONTROL
   "Carrier_78_G120DControlWord.0" AT %I4260.0 : Bool;   // Bit_00_ON
   "Carrier_78_G120DControlWord.1" AT %I4260.1 : Bool;   // Bit_01_AUS2_INH
   "Carrier_78_G120DControlWord.2" AT %I4260.2 : Bool;   // Bit_02_AUS3_STOP
   "Carrier_78_G120DControlWord.3" AT %I4260.3 : Bool;   // Bit_03_EN
   "Carrier_78_G120DControlWord.4" AT %I4260.4 : Bool;   // Bit_04_EN_RAMP
   "Carrier_78_G120DControlWord.5" AT %I4260.5 : Bool;   // Bit_05_START_RAMP
   "Carrier_78_G120DControlWord.6" AT %I4260.6 : Bool;   // Bit_06_SETPOINT
   "Carrier_78_G120DControlWord.7" AT %I4260.7 : Bool;   // Bit_07_RESET
   "Carrier_78_G120DControlWord.8" AT %I4261.0 : Bool;   // Bit_08_JOG_R
   "Carrier_78_G120DControlWord.9" AT %I4261.1 : Bool;   // Bit_09_JOG_L
   "Carrier_78_G120DControlWord.10" AT %I4261.2 : Bool;   // Bit_10_CONTR_PLC
   "Carrier_78_G120DControlWord.11" AT %I4261.3 : Bool;   // Bit_11_REVERSE
   "Carrier_78_G120DControlWord.12" AT %I4261.4 : Bool;   // Bit_12_BRAKE_RELEASE
   "Carrier_78_G120DControlWord.13" AT %I4261.5 : Bool;   // Bit_13_DDS
   "Carrier_78_G120DControlWord.14" AT %I4261.6 : Bool;   // Bit_14_DO0
   "Carrier_78_G120DControlWord.15" AT %I4261.7 : Bool;   // Bit_15_DO1
   "Carrier_78_G120DStatusWord" AT %IW4262 : Word;   // G120D_ZSW1_STATUS
   "Carrier_78_G120DStatusWord.0" AT %I4262.0 : Bool;   // Bit_00_READY_RUN
   "Carrier_78_G120DStatusWord.1" AT %I4262.1 : Bool;   // Bit_01_READY_ON
   "Carrier_78_G120DStatusWord.2" AT %I4262.2 : Bool;   // Bit_02_ENABLE
   "Carrier_78_G120DStatusWord.3" AT %I4262.3 : Bool;   // Bit_03_FAULT
   "Carrier_78_G120DStatusWord.4" AT %I4262.4 : Bool;   // Bit_04_OFF2
   "Carrier_78_G120DStatusWord.5" AT %I4262.5 : Bool;   // Bit_05_OFF3
   "Carrier_78_G120DStatusWord.6" AT %I4262.6 : Bool;   // Bit_06_LOCK_OUT
   "Carrier_78_G120DStatusWord.7" AT %I4262.7 : Bool;   // Bit_07_WARN
   "Carrier_78_G120DStatusWord.8" AT %I4263.0 : Bool;   // Bit_08_NO_DEVIATION
   "Carrier_78_G120DStatusWord.9" AT %I4263.1 : Bool;   // Bit_09_CONTR_PLC
   "Carrier_78_G120DStatusWord.10" AT %I4263.2 : Bool;   // Bit_10_F_MAX
   "Carrier_78_G120DStatusWord.11" AT %I4263.3 : Bool;   // Bit_11_LIMIT_REACHED
   "Carrier_78_G120DStatusWord.12" AT %I4263.4 : Bool;   // Bit_12_BRAKE_OPEN
   "Carrier_78_G120DStatusWord.13" AT %I4263.5 : Bool;   // Bit_13_NO_OVERTEMP
   "Carrier_78_G120DStatusWord.14" AT %I4263.6 : Bool;   // Bit_14_CW_CCW
   "Carrier_78_G120DStatusWord.15" AT %I4263.7 : Bool;   // Bit_15_OVERL
   "Carrier_78_Slot2_Input" AT %IW4264 : Word;   // SLOT 2 INPUT WORD
   "Carrier_78_CrashDetectSW" AT %I4264.0 : Bool;   // CRASH DETECT SW
   "Carrier_78_SpareSafetyInput(2_1)" AT %I4264.1 : Bool;   // SPARE SAFETY INPUT
   "Carrier_78_SpareSafetyInput(2_2)" AT %I4264.2 : Bool;   // SPARE SAFETY INPUT